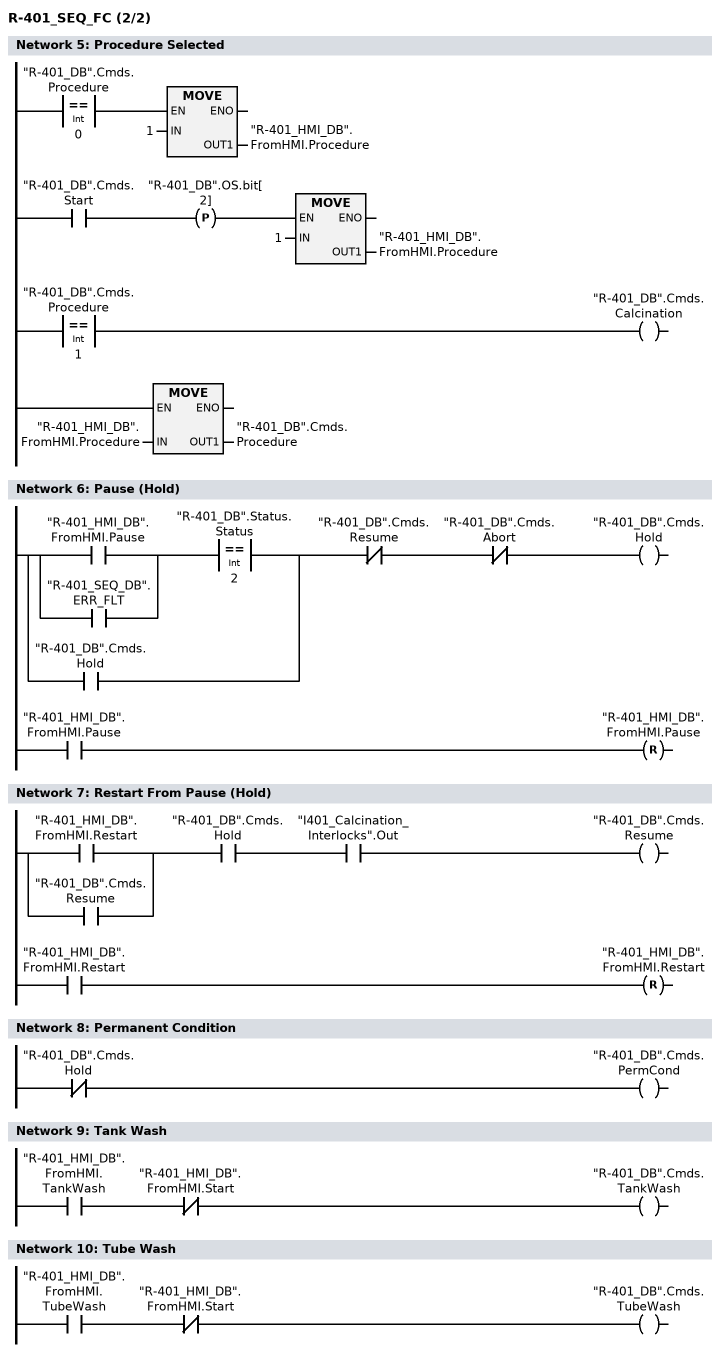
   RUNG wire#powerrail
      { S7_Templates := "SrcType := Int" } EQ_Contact(in1 := "R-401_DB".Cmds.Procedure, in2 := 0)
      Move(in := 1, out1 => "R-401_HMI_DB".FromHMI.Procedure)
   END_RUNG
   RUNG wire#powerrail
      Contact( "R-401_DB".Cmds.Start )
      P_Trig( "R-401_DB".OS.bit[2] )
      Move(in := 1, out1 => "R-401_HMI_DB".FromHMI.Procedure)
   END_RUNG
   RUNG wire#powerrail
      { S7_Templates := "SrcType := Int" } EQ_Contact(in1 := "R-401_DB".Cmds.Procedure, in2 := 1)
      Coil( "R-401_DB".Cmds.Calcination )
   END_RUNG
   RUNG wire#powerrail
      Move(in := "R-401_HMI_DB".FromHMI.Procedure, out1 => "R-401_DB".Cmds.Procedure)
   END_RUNG
   // the same network as SCL:
   IF "R-401_DB".Cmds.Procedure = 0 THEN "R-401_HMI_DB".FromHMI.Procedure := 1; END_IF;
   #_w1 := "R-401_DB".Cmds.Start AND NOT "R-401_DB".OS.bit[2];   // rising edge
   "R-401_DB".OS.bit[2] := "R-401_DB".Cmds.Start;
   IF #_w1 THEN "R-401_HMI_DB".FromHMI.Procedure := 1; END_IF;
   "R-401_DB".Cmds.Calcination := "R-401_DB".Cmds.Procedure = 1;
   "R-401_DB".Cmds.Procedure := "R-401_HMI_DB".FromHMI.Procedure;
END_REGION

REGION Network 6: Pause (Hold)
   RUNG wire#powerrail
      Contact( "R-401_HMI_DB".FromHMI.Pause )
      wire#w1
      { S7_Templates := "SrcType := Int" } EQ_Contact(in1 := "R-401_DB".Status.Status, in2 := 2)
      wire#w2
      I_Contact( "R-401_DB".Cmds.Resume )
      I_Contact( "R-401_DB".Cmds.Abort )
      Coil( "R-401_DB".Cmds.Hold )
   END_RUNG
   RUNG wire#powerrail
      Contact( "R-401_SEQ_DB".ERR_FLT )
   END_RUNG wire#w1
   RUNG wire#powerrail
      Contact( "R-401_DB".Cmds.Hold )
   END_RUNG wire#w2
   RUNG wire#powerrail
      Contact( "R-401_HMI_DB".FromHMI.Pause )
      R_Coil( "R-401_HMI_DB".FromHMI.Pause )
   END_RUNG
   // the same network as SCL:
   "R-401_DB".Cmds.Hold := ((("R-401_HMI_DB".FromHMI.Pause OR "R-401_SEQ_DB".ERR_FLT) AND ("R-401_DB".Status.Status = 2)) OR "R-401_DB".Cmds.Hold) AND NOT "R-401_DB".Cmds.Resume AND NOT "R-401_DB".Cmds.Abort;
   IF "R-401_HMI_DB".FromHMI.Pause THEN "R-401_HMI_DB".FromHMI.Pause := FALSE; END_IF;
END_REGION

REGION Network 7: Restart From Pause (Hold)
   RUNG wire#powerrail
      Contact( "R-401_HMI_DB".FromHMI.Restart )
      wire#w1
      Contact( "R-401_DB".Cmds.Hold )
      Contact( "I401_Calcination_Interlocks".Out )
      Coil( "R-401_DB".Cmds.Resume )
   END_RUNG
   RUNG wire#powerrail
      Contact( "R-401_DB".Cmds.Resume )
   END_RUNG wire#w1
   RUNG wire#powerrail
      Contact( "R-401_HMI_DB".FromHMI.Restart )
      R_Coil( "R-401_HMI_DB".FromHMI.Restart )
   END_RUNG
   // the same network as SCL:
   "R-401_DB".Cmds.Resume := ("R-401_HMI_DB".FromHMI.Restart OR "R-401_DB".Cmds.Resume) AND "R-401_DB".Cmds.Hold AND "I401_Calcination_Interlocks".Out;
   IF "R-401_HMI_DB".FromHMI.Restart THEN "R-401_HMI_DB".FromHMI.Restart := FALSE; END_IF;
END_REGION

REGION Network 8: Permanent Condition
   RUNG wire#powerrail
      I_Contact( "R-401_DB".Cmds.Hold )
      Coil( "R-401_DB".Cmds.PermCond )
   END_RUNG
   // the same network as SCL:
   "R-401_DB".Cmds.PermCond := NOT "R-401_DB".Cmds.Hold;
END_REGION

REGION Network 9: Tank Wash
   RUNG wire#powerrail
      Contact( "R-401_HMI_DB".FromHMI.TankWash )
      I_Contact( "R-401_HMI_DB".FromHMI.Start )
      Coil( "R-401_DB".Cmds.TankWash )
   END_RUNG
   // the same network as SCL:
   "R-401_DB".Cmds.TankWash := "R-401_HMI_DB".FromHMI.TankWash AND NOT "R-401_HMI_DB".FromHMI.Start;
END_REGION

REGION Network 10: Tube Wash
   RUNG wire#powerrail
      Contact( "R-401_HMI_DB".FromHMI.TubeWash )
      I_Contact( "R-401_HMI_DB".FromHMI.Start )
      Coil( "R-401_DB".Cmds.TubeWash )
   END_RUNG
   // the same network as SCL:
   "R-401_DB".Cmds.TubeWash := "R-401_HMI_DB".FromHMI.TubeWash AND NOT "R-401_HMI_DB".FromHMI.Start;
END_REGION

REGION Network 11 (SCL): Sequence Status
   IF "R-401_SEQ_DB".S_NO= 1 THEN
       "R-401_DB".Status.Status := 1; //Idle
   ELSIF (("R-401_SEQ_DB".S_NO > 1 AND "R-401_SEQ_DB".S_NO < 150) OR ("R-401_SEQ_DB".S_NO > 161 AND "R-401_SEQ_DB".S_NO < 170)) AND NOT "R-401_SEQ_DB".ERR_FLT AND NOT "R-401_DB".Cmds.Hold THEN
       "R-401_DB".Status.Status := 2; //Running
   ELSIF "R-401_SEQ_DB".S_NO >= 151 AND "R-401_SEQ_DB".S_NO <= 160 AND NOT "R-401_SEQ_DB".ERR_FLT THEN
       "R-401_DB".Status.Status := 3; // Stopping
   ELSIF  "R-401_SEQ_DB".ERR_FLT AND  (("R-401_SEQ_DB".S_NO > 1 AND "R-401_SEQ_DB".S_NO < 150) OR ("R-401_SEQ_DB".S_NO > 161 AND "R-401_SEQ_DB".S_NO < 170)) THEN
       "R-401_DB".Status.Status := 4; // Held
   ELSIF  "R-401_SEQ_DB".ERR_FLT AND  (("R-401_SEQ_DB".S_NO > 1 AND "R-401_SEQ_DB".S_NO < 150) OR ("R-401_SEQ_DB".S_NO > 161 AND "R-401_SEQ_DB".S_NO < 170)) AND "R-401_Aux_DB"."Bool".TOff  THEN
       "R-401_DB".Status.Status := 5; // Holding
   ELSE
       "R-401_DB".Status.Status := 6; // Unknown
   END_IF;

   "R-401_DB".Status.Running := ("R-401_SEQ_DB".S_NO > 3 AND "R-401_SEQ_DB".S_NO < 150) OR ("R-401_SEQ_DB".S_NO > 161 AND "R-401_SEQ_DB".S_NO < 170);
   "R-401_DB".Status.Initializing := ("R-401_SEQ_DB".S_NO >= 141 AND "R-401_SEQ_DB".S_NO <= 150);

   //Enable/Disable HMI Start/Stop Button
   "R-401_HMI_DB".ToHMI.EnStopButton := ("R-401_DB".Status.Status > 1) OR "R-401_DB".Status.Step = 0; //Enable HMI Stop Button
   "R-401_HMI_DB".ToHMI.EnStartButton := "R-401_DB".Status.Status = 1; //Idle
   "R-401_HMI_DB".ToHMI.EnPauseButton := "R-401_DB".Status.Status = 2; //Enable Pause Button
   "R-401_HMI_DB".ToHMI.EnRestartButton :=  "R-401_DB".Status.Status = 4; //Enable Restart Button

   //****Interlock Activated
   "R-401_HMI_DB".ToHMI.InterlockActivated := "I401_Calcination_Interlocks".Out;
END_REGION

REGION Network 12 (SCL): Sequence Step
   "R-401_DB".Status.Step := "R-401_SEQ_DB".S_NO;
END_REGION

REGION Network 13 (SCL): Sequence state (Procedure running)
   IF "R-401_SEQ_DB".S_NO = 3 OR "R-401_SEQ_DB".S_NO = 4 THEN
       "R-401_DB".Status.State := 1; //Ready
   ELSIF "R-401_SEQ_DB".S_NO >= 21 AND "R-401_SEQ_DB".S_NO <= 60 THEN
       "R-401_DB".Status.State := 2; //Mixing 
   ELSIF "R-401_SEQ_DB".S_NO >= 61 AND "R-401_SEQ_DB".S_NO <= 80 THEN
       "R-401_DB".Status.State := 3; //Pouring
   ELSIF "R-401_SEQ_DB".S_NO >= 141 AND "R-401_SEQ_DB".S_NO <= 150 THEN
       "R-401_DB".Status.State := 4; //Initializing
   ELSIF "R-401_SEQ_DB".S_NO >= 151 AND "R-401_SEQ_DB".S_NO <= 160 THEN
       "R-401_DB".Status.State := 5; //Aborting
   ELSE
       "R-401_DB".Status.State := 0;
   END_IF;
END_REGION

REGION Network 14: Sequence State
END_REGION
END_FUNCTION

FUNCTION "R-401_Tansitions_FC" : Void   // FC98, SCL
{ S7_Optimized_Access := 'TRUE' }
VERSION : 0.1
   VAR_TEMP
      Cond : Struct
         CtrlsOff : Bool;
         Steps : Bool;
      END_STRUCT;
   END_VAR
BEGIN


   //********Controllers Off********
   #Cond.CtrlsOff:= "TC-4011A_R3".MB_Data.Buffer[1] = 0 AND "TC-4011A_R3".MB_Data.Buffer[1] = 0 AND "TC-4011A_R3".MB_Data.Buffer[1] = 0;
   //********Steps********
   #Cond.Steps := "R-401_DB".Status.Step = 25 OR "R-401_DB".Status.Step = 27 OR "R-401_DB".Status.Step = 29;

   //*****************************************Transition conditions**************************************

   "R-401_Aux_DB"."Bool".Cond._001 := #Cond.CtrlsOff;      //"R401_TempMon_DB".ReadyToProcess  AND
END_FUNCTION

// folder: State MACHINE/5)Passivate

FUNCTION "Monitor_R402_FC" : Void   // FC99, LAD
TITLE = FC to call User Functions
{ S7_Optimized_Access := 'TRUE' }
AUTHOR : JL
VERSION : 0.1
BEGIN

REGION Network 1: Moving Furnace temperature to the monitor block
   // Thermocouples:
   // "TT-401A_DB".SAI
   // "TT-401B_DB".SAI
   // "TT-401C_DB".SAI
   // "TT-401C_DB".SAI
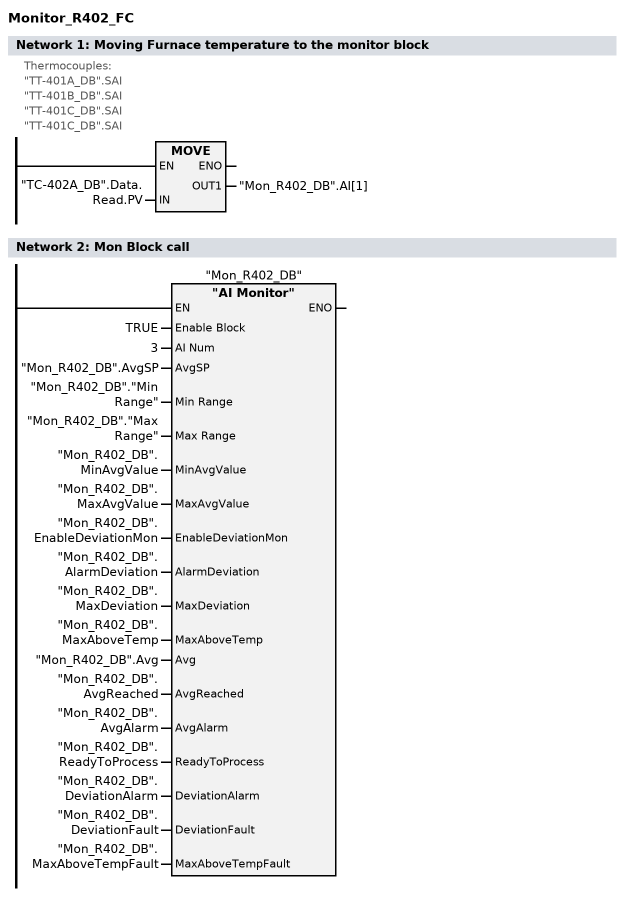
   RUNG wire#powerrail
      Move(in := "TC-402A_DB".Data.Read.PV, out1 => "Mon_R402_DB".AI[1])
   END_RUNG
   // the same network as SCL:
   "Mon_R402_DB".AI[1] := "TC-402A_DB".Data.Read.PV;
END_REGION

REGION Network 2: Mon Block call
   RUNG wire#powerrail
      "Mon_R402_DB"("Enable Block" := TRUE, "AI Num" := 3, AvgSP := "Mon_R402_DB".AvgSP, "Min Range" := "Mon_R402_DB"."Min Range", "Max Range" := "Mon_R402_DB"."Max Range", MinAvgValue := "Mon_R402_DB".MinAvgValue, MaxAvgValue := "Mon_R402_DB".MaxAvgValue, EnableDeviationMon := "Mon_R402_DB".EnableDeviationMon, AlarmDeviation := "Mon_R402_DB".AlarmDeviation, MaxDeviation := "Mon_R402_DB".MaxDeviation, MaxAboveTemp := "Mon_R402_DB".MaxAboveTemp, Avg := "Mon_R402_DB".Avg, AvgReached := "Mon_R402_DB".AvgReached, AvgAlarm := "Mon_R402_DB".AvgAlarm, ReadyToProcess := "Mon_R402_DB".ReadyToProcess, DeviationAlarm := "Mon_R402_DB".DeviationAlarm, DeviationFault := "Mon_R402_DB".DeviationFault, MaxAboveTempFault := "Mon_R402_DB".MaxAboveTempFault)
   END_RUNG
   // the same network as SCL:
   "Mon_R402_DB"("Enable Block" := TRUE,   // "AI Monitor"
                 "AI Num" := 3,
                 AvgSP := "Mon_R402_DB".AvgSP,
                 "Min Range" := "Mon_R402_DB"."Min Range",
                 "Max Range" := "Mon_R402_DB"."Max Range",
                 MinAvgValue := "Mon_R402_DB".MinAvgValue,
                 MaxAvgValue := "Mon_R402_DB".MaxAvgValue,
                 EnableDeviationMon := "Mon_R402_DB".EnableDeviationMon,
                 AlarmDeviation := "Mon_R402_DB".AlarmDeviation,
                 MaxDeviation := "Mon_R402_DB".MaxDeviation,
                 MaxAboveTemp := "Mon_R402_DB".MaxAboveTemp,
                 Avg := "Mon_R402_DB".Avg,
                 AvgReached := "Mon_R402_DB".AvgReached,
                 AvgAlarm := "Mon_R402_DB".AvgAlarm,
                 ReadyToProcess := "Mon_R402_DB".ReadyToProcess,
                 DeviationAlarm := "Mon_R402_DB".DeviationAlarm,
                 DeviationFault := "Mon_R402_DB".DeviationFault,
                 MaxAboveTempFault := "Mon_R402_DB".MaxAboveTempFault);
END_REGION
END_FUNCTION

// folder: State MACHINE/5)Passivate/Reactor R-402

FUNCTION_BLOCK "R-402_SEQ"   // FB31, GRAPH_PLUS
TITLE = Reactor R-401
{ S7_Optimized_Access := 'TRUE' }
AUTHOR : JL
VERSION : 0.1
   VAR_INPUT
      OFF_SQ : Bool := false;   // Turn sequence off
      INIT_SQ : Bool := false;   // Set sequence to initial state
      ACK_EF : Bool := false;   // Acknowledge all errors and faults
      S_PREV : Bool := false;   // Output previous step in parameter S_NO
      S_NEXT : Bool := false;   // Indicate next step in parameter S_NO
      SW_AUTO : Bool := false;   // Automatic mode
      SW_TAP : Bool := false;   // Semiautomatic/switch with transition
      SW_TOP : Bool := false;   // Semiautomatic/ignore transition
      SW_MAN : Bool := false;   // Manual mode
      S_SEL : Int := 0;   // Select step to be output to S_NO
      S_ON : Bool := false;   // Activate step indicated in S_NO
      S_OFF : Bool := false;   // Deactivate step indicated S_NO
      T_PUSH : Bool := false;   // Enable transition to switch in semi automatic mode
   END_VAR
   VAR_OUTPUT
      S_NO : Int := 0;   // Step number
      S_MORE : Bool := false;   // More steps are available and can be shown in S_NO
      S_ACTIVE : Bool := false;   // Step indicated in S_NO is active
      ERR_FLT : Bool := false;   // Interlock or supervision group error
      AUTO_ON : Bool := false;   // Automatic mode is active
      TAP_ON : Bool := false;   // Semiautomatic mode/step with transition enabled
      TOP_ON : Bool := false;   // Semiautomatic mode/ignore transition enabled
      MAN_ON : Bool := false;   // Manual mode is active
   END_VAR
   VAR
      HMI_INFO : Array[0..12] of UInt;
      IF_PAR : G7_IfParPlus_V6;
      RT_DATA : G7_RTDataPlus_V6;   // Internal data area
      Abort : G7_TransitionPlus_V6;   // Transition structure
      InitializeR : G7_TransitionPlus_V6;   // Transition structure
      CalcinP : G7_TransitionPlus_V6;   // Transition structure
      Re : G7_TransitionPlus_V6;   // Transition structure
      Calcinat : G7_TransitionPlus_V6;   // Transition structure
      Wash : G7_TransitionPlus_V6;   // Transition structure
      Shutdwn : G7_TransitionPlus_V6;   // Transition structure
      ColdDDn : G7_TransitionPlus_V6;   // Transition structure
      Std : G7_TransitionPlus_V6;   // Transition structure
      PDn : G7_TransitionPlus_V6;   // Transition structure
      PressRd : G7_TransitionPlus_V6;   // Transition structure
      Rmp1Dn : G7_TransitionPlus_V6;   // Transition structure
      FHldDn : G7_TransitionPlus_V6;   // Transition structure
      Rmp2Dn : G7_TransitionPlus_V6;   // Transition structure
      ScHldDn : G7_TransitionPlus_V6;   // Transition structure
      Rmp3Dn : G7_TransitionPlus_V6;   // Transition structure
      ThHldDn : G7_TransitionPlus_V6;   // Transition structure
      Trans30 : G7_TransitionPlus_V6;   // Transition structure
      Trans31 : G7_TransitionPlus_V6;   // Transition structure
      End : G7_TransitionPlus_V6;   // Transition structure
      Init : G7_TransitionPlus_V6;   // Transition structure
      SAut : G7_TransitionPlus_V6;   // Transition structure
      SIn : G7_TransitionPlus_V6;   // Transition structure
      Initd : G7_TransitionPlus_V6;   // Transition structure
      Ab : G7_TransitionPlus_V6;   // Transition structure
      AbortOn : G7_TransitionPlus_V6;   // Transition structure
      AbortDn : G7_TransitionPlus_V6;   // Transition structure
      ShtSted : G7_TransitionPlus_V6;   // Transition structure
      CldDwnDn : G7_TransitionPlus_V6;   // Transition structure
      DPDn : G7_TransitionPlus_V6;   // Transition structure
      Idle : G7_StepPlus_V6;   // Step structure
      Ready : G7_StepPlus_V6;   // Step structure
      SelectSeq : G7_StepPlus_V6;   // Step structure
      Started : G7_StepPlus_V6;   // Step structure
      "EDIT Params" : G7_StepPlus_V6;   // Step structure
      "USER StartN2" : G7_StepPlus_V6;   // Step structure
      RampUp1 : G7_StepPlus_V6;   // Step structure
      CloseN2 : G7_StepPlus_V6;   // Step structure
      HoldTime : G7_StepPlus_V6;   // Step structure
      SecondHold : G7_StepPlus_V6;   // Step structure
      RampUp3 : G7_StepPlus_V6;   // Step structure
      ThirdHold : G7_StepPlus_V6;   // Step structure
      HeatersOff : G7_StepPlus_V6;   // Step structure
      PressureOff : G7_StepPlus_V6;   // Step structure
      Done : G7_StepPlus_V6;   // Step structure
      Initialize : G7_StepPlus_V6;   // Step structure
      SetAuto : G7_StepPlus_V6;   // Step structure
      SetInitial : G7_StepPlus_V6;   // Step structure
      Initialized : G7_StepPlus_V6;   // Step structure
      AbortStarting : G7_StepPlus_V6;   // Step structure
      Aborting : G7_StepPlus_V6;   // Step structure
      AbortDone : G7_StepPlus_V6;   // Step structure
      ShtdnStarted : G7_StepPlus_V6;   // Step structure
      CoolingDown : G7_StepPlus_V6;   // Step structure
      DePress : G7_StepPlus_V6;   // Step structure
      ShtdnDn : G7_StepPlus_V6;   // Step structure
      SINI : Array[0..5] of USInt;
      LSTT : Array[0..29] of USInt;
      ATAJ : Array[0..29] of USInt;
      ATAB : Array[0..29] of USInt;
      PSTT : Array[0..29] of USInt;
      NSTT : Array[0..29] of USInt;
      ASSJ : Array[0..25] of USInt;
      ASSB : Array[0..25] of USInt;
      PTTS : Array[0..25] of USInt;
      NTTS : Array[0..25] of USInt;
      SW_SQTS : Array[0..25] of USInt;
      SWITCH : Array[0..4] of USInt;
      TVX : Array[0..11] of USInt;
      TTX : Array[0..11] of USInt;
      TSX : Array[0..5] of USInt;
      S00X : Array[0..5] of USInt;
      SOFFX : Array[0..5] of USInt;
      SONX : Array[0..5] of USInt;
      SAX : Array[0..5] of USInt;
      SERRX : Array[0..26] of USInt;
      SMX : Array[0..26] of USInt;
      S0X : Array[0..26] of USInt;
      S1X : Array[0..26] of USInt;
      IL_ALARM_INST : Diag_Alarm;
      SUP_ALARM_INST : Diag_Alarm;
      STEP_TIME_ALARM_INST : Diag_Alarm;
      IEC_TIMER_INST : IEC_TIMER;
      TRANSACTION_FLAG : Bool := false;
   END_VAR
   // SINI[0] := 2;
   // LSTT[0] := 19;
   // NSTT[0] := 19;
   // PTTS[0] := 255;
   // TVX[0] := 16#1;
   // TTX[0] := 16#1;
   // TSX[0] := 16#1;
   // S00X[0] := 16#1;
   // SOFFX[0] := 16#1;
   // SONX[0] := 16#1;
   // SAX[0] := 16#1;
   // SERRX[0] := 16#1;
   // SMX[0] := 16#1;
   // S0X[0] := 16#1;
   // S1X[0] := 16#1;
   // SINI[2] := 255;
   // SINI[3] := 255;
   // SINI[4] := 255;
   // LSTT[1] := 15;
   // LSTT[2] := 255;
   // LSTT[3] := 255;
   // LSTT[4] := 3;
   // LSTT[5] := 255;
   // LSTT[6] := 22;
   // LSTT[16] := 255;
   // LSTT[8] := 255;
   // LSTT[9] := 255;
   // LSTT[10] := 255;
   // LSTT[11] := 255;
   // LSTT[12] := 255;
   // LSTT[13] := 255;
   // LSTT[14] := 255;
   // LSTT[19] := 255;
   // LSTT[22] := 255;
   // LSTT[17] := 255;
   // LSTT[25] := 255;
   // LSTT[20] := 255;
   // LSTT[21] := 255;
   // ATAJ[1] := 1;
   // ATAJ[2] := 2;
   // ATAJ[3] := 3;
   // ATAJ[4] := 4;
   // ATAJ[5] := 5;
   // ATAJ[6] := 6;
   // ATAJ[7] := 7;
   // ATAJ[8] := 8;
   // ATAJ[9] := 9;
   // ATAJ[10] := 10;
   // ATAJ[11] := 11;
   // ATAJ[12] := 12;
   // ATAJ[13] := 13;
   // ATAJ[14] := 14;
   // ATAJ[15] := 15;
   // ATAJ[16] := 16;
   // ATAJ[17] := 17;
   // ATAJ[18] := 18;
   // ATAJ[19] := 19;
   // ATAJ[20] := 20;
   // ATAJ[21] := 21;
   // ATAJ[22] := 22;
   // ATAB[0] := 6;
   // ATAB[1] := 2;
   // ATAB[3] := 3;
   // ATAB[4] := 5;
   // ATAB[5] := 4;
   // ATAB[6] := 1;
   // ATAB[7] := 7;
   // ATAB[8] := 8;
   // ATAB[9] := 9;
   // ATAB[10] := 10;
   // ATAB[11] := 11;
   // ATAB[12] := 12;
   // ATAB[13] := 13;
   // ATAB[14] := 14;
   // ATAB[15] := 15;
   // ATAB[16] := 16;
   // ATAB[17] := 17;
   // ATAB[18] := 18;
   // ATAB[19] := 19;
   // ATAB[20] := 20;
   // ATAB[21] := 21;
   // ATAB[22] := 22;
   // SW_SQTS[21] := 4;
   // SW_SQTS[20] := 4;
   // PSTT[3] := 1;
   // PSTT[4] := 2;
   // PSTT[5] := 2;
   // PSTT[22] := 17;
   // PSTT[7] := 25;
   // PSTT[8] := 3;
   // PSTT[9] := 4;
   // PSTT[10] := 5;
   // PSTT[11] := 6;
   // PSTT[12] := 7;
   // PSTT[13] := 8;
   // PSTT[14] := 9;
   // PSTT[15] := 10;
   // PSTT[16] := 11;
   // PSTT[17] := 13;
   // PSTT[18] := 14;
   // PSTT[19] := 12;
   // PSTT[20] := 15;
   // PSTT[21] := 16;
   // PSTT[25] := 20;
   // NTTS[21] := 26;
   // NTTS[20] := 25;
   // PTTS[21] := 25;
   // PTTS[20] := 24;
   // NSTT[1] := 15;
   // NSTT[2] := 1;
   // NSTT[3] := 2;
   // NSTT[4] := 3;
   // NSTT[5] := 255;
   // NSTT[6] := 22;
   // NSTT[16] := 12;
   // NSTT[8] := 4;
   // NSTT[9] := 5;
   // NSTT[10] := 6;
   // NSTT[11] := 7;
   // NSTT[12] := 8;
   // NSTT[13] := 9;
   // NSTT[14] := 10;
   // NSTT[19] := 13;
   // NSTT[22] := 18;
   // NSTT[17] := 14;
   // NSTT[25] := 21;
   // NSTT[20] := 16;
   // NSTT[21] := 17;
   // ASSJ[20] := 20;
   // ASSB[21] := 21;
   // ASSB[20] := 20;
   // ASSJ[21] := 21;
   // ASSJ[1] := 1;
   // ASSJ[2] := 2;
   // ASSJ[3] := 3;
   // ASSJ[4] := 4;
   // ASSJ[5] := 5;
   // ASSJ[6] := 6;
   // ASSJ[7] := 7;
   // ASSJ[8] := 8;
   // ASSJ[9] := 9;
   // ASSJ[10] := 10;
   // ASSJ[11] := 11;
   // ASSJ[12] := 12;
   // ASSJ[13] := 13;
   // ASSJ[14] := 14;
   // ASSJ[15] := 15;
   // ASSJ[16] := 16;
   // ASSJ[17] := 17;
   // ASSJ[18] := 18;
   // ASSJ[19] := 19;
   // NSTT[23] := 1;
   // NSTT[15] := 11;
   // PSTT[24] := 19;
   // PSTT[23] := 18;
   // ASSB[1] := 1;
   // ASSB[2] := 2;
   // ASSB[3] := 3;
   // ASSB[4] := 4;
   // ASSB[5] := 5;
   // ASSB[6] := 6;
   // ASSB[7] := 7;
   // ASSB[8] := 8;
   // ASSB[9] := 9;
   // ASSB[10] := 10;
   // ASSB[11] := 11;
   // ASSB[12] := 12;
   // ASSB[13] := 13;
   // ASSB[14] := 14;
   // ASSB[15] := 15;
   // ASSB[16] := 16;
   // ASSB[17] := 17;
   // ASSB[18] := 18;
   // ASSB[19] := 19;
   // ATAB[24] := 24;
   // ATAB[23] := 23;
   // ATAJ[24] := 24;
   // ATAJ[23] := 23;
   // PTTS[1] := 2;
   // PTTS[2] := 3;
   // PTTS[3] := 255;
   // PTTS[4] := 8;
   // PTTS[5] := 9;
   // PTTS[6] := 10;
   // PTTS[7] := 11;
   // PTTS[8] := 12;
   // PTTS[9] := 13;
   // PTTS[10] := 14;
   // PTTS[11] := 15;
   // PTTS[12] := 16;
   // PTTS[13] := 19;
   // PTTS[14] := 17;
   // PTTS[15] := 255;
   // PTTS[16] := 20;
   // PTTS[17] := 21;
   // PTTS[18] := 22;
   // PTTS[19] := 255;
   // LSTT[23] := 1;
   // LSTT[15] := 255;
   // NTTS[1] := 3;
   // NTTS[2] := 4;
   // NTTS[3] := 8;
   // NTTS[4] := 9;
   // NTTS[5] := 10;
   // NTTS[6] := 11;
   // NTTS[7] := 12;
   // NTTS[8] := 13;
   // NTTS[9] := 14;
   // NTTS[10] := 15;
   // NTTS[11] := 16;
   // NTTS[12] := 19;
   // NTTS[13] := 17;
   // NTTS[14] := 18;
   // NTTS[15] := 20;
   // NTTS[16] := 21;
   // NTTS[17] := 22;
   // NTTS[18] := 23;
   // NTTS[19] := 24;
   // SW_SQTS[1] := 1;
   // SW_SQTS[2] := 1;
   // SW_SQTS[3] := 2;
   // SW_SQTS[4] := 2;
   // SW_SQTS[5] := 2;
   // SW_SQTS[6] := 2;
   // SW_SQTS[7] := 2;
   // SW_SQTS[8] := 2;
   // SW_SQTS[9] := 2;
   // SW_SQTS[10] := 2;
   // SW_SQTS[11] := 2;
   // SW_SQTS[12] := 2;
   // SW_SQTS[13] := 2;
   // SW_SQTS[14] := 2;
   // SW_SQTS[15] := 3;
   // SW_SQTS[16] := 3;
   // SW_SQTS[17] := 3;
   // SW_SQTS[18] := 3;
   // SW_SQTS[19] := 4;
   // SWITCH[0] := 60;
   // SWITCH[1] := 191;
   // SWITCH[2] := 223;
   // SINI[5] := 255;
   // LSTT[24] := 255;
   // LSTT[28] := 255;
   // LSTT[27] := 255;
   // ATAJ[25] := 25;
   // ATAJ[26] := 26;
   // ATAJ[27] := 27;
   // ATAJ[28] := 28;
   // ATAB[25] := 25;
   // ATAB[26] := 26;
   // ATAB[27] := 27;
   // ATAB[28] := 28;
   // PSTT[26] := 21;
   // PSTT[27] := 22;
   // PSTT[28] := 23;
   // NSTT[24] := 20;
   // NSTT[28] := 24;
   // NSTT[27] := 23;
   // ASSJ[22] := 22;
   // ASSJ[23] := 23;
   // ASSJ[24] := 24;
   // ASSB[22] := 22;
   // ASSB[23] := 23;
   // ASSB[24] := 24;
   // PTTS[22] := 255;
   // PTTS[23] := 27;
   // PTTS[24] := 28;
   // NTTS[22] := 27;
   // NTTS[23] := 28;
   // NTTS[24] := 29;
   // SW_SQTS[22] := 5;
   // SW_SQTS[23] := 5;
   // SW_SQTS[24] := 5;
   // SWITCH[3] := 239;
   // SWITCH[4] := 7;
   // LSTT[29] := 255;
   // ATAJ[29] := 29;
   // ATAB[29] := 29;
   // PSTT[29] := 24;
   // NSTT[29] := 25;
   // ASSJ[25] := 25;
   // ASSB[25] := 25;
   // PTTS[25] := 29;
   // NTTS[25] := 7;
   // SW_SQTS[25] := 5;
BEGIN
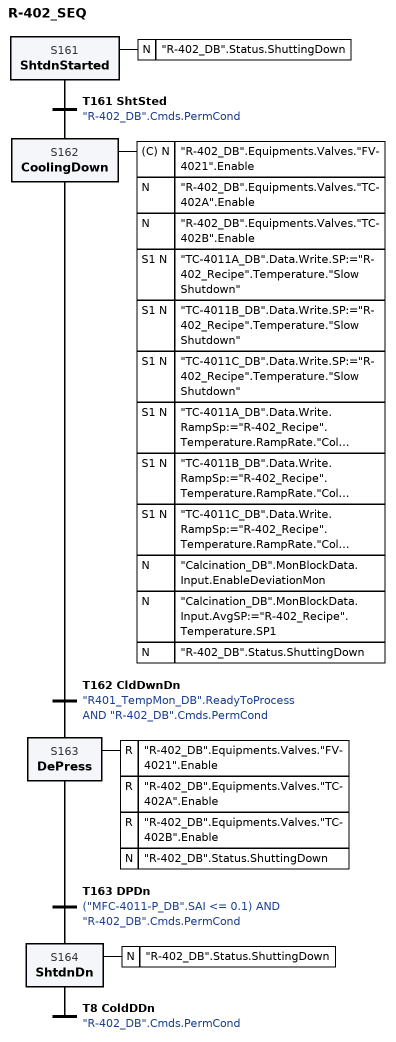
   // permanent pre-instructions
   NETWORK 1
      "R-402_SEQ_FC"();
      "R-402_FC_Inputs"();
      "Monitor_R402_FC"();
      "Alarms"();

   // sequencer 1
   STEP ShtdnStarted:   // S161, max time T#10S, warning time T#7S
      // Shutdown Started
              N    "R-402_DB".Status.ShuttingDown
   END_STEP
   TRANSITION ShtSted FROM ShtdnStarted TO CoolingDown   // T161
      := "R-402_DB".Cmds.PermCond;
   END_TRANSITION
   STEP CoolingDown:   // S162, max time T#10S, warning time T#7S
      (C)     N    "R-402_DB".Equipments.Valves."FV-4021".Enable
              N    "R-402_DB".Equipments.Valves."TC-402A".Enable
              N    "R-402_DB".Equipments.Valves."TC-402B".Enable
          S1  N    "TC-4011A_DB".Data.Write.SP:="R-402_Recipe".Temperature."Slow Shutdown"
          S1  N    "TC-4011B_DB".Data.Write.SP:="R-402_Recipe".Temperature."Slow Shutdown"
          S1  N    "TC-4011C_DB".Data.Write.SP:="R-402_Recipe".Temperature."Slow Shutdown"
          S1  N    "TC-4011A_DB".Data.Write.RampSp:="R-402_Recipe".Temperature.RampRate."Cold Down"
          S1  N    "TC-4011B_DB".Data.Write.RampSp:="R-402_Recipe".Temperature.RampRate."Cold Down"
          S1  N    "TC-4011C_DB".Data.Write.RampSp:="R-402_Recipe".Temperature.RampRate."Cold Down"
              N    "Calcination_DB".MonBlockData.Input.EnableDeviationMon
              N    "Calcination_DB".MonBlockData.Input.AvgSP:="R-402_Recipe".Temperature.SP1
              N    "R-402_DB".Status.ShuttingDown
   END_STEP
   TRANSITION CldDwnDn FROM CoolingDown TO DePress   // T162
      := "R401_TempMon_DB".ReadyToProcess AND "R-402_DB".Cmds.PermCond;
   END_TRANSITION
   STEP DePress:   // S163, max time T#10S, warning time T#7S
              R    "R-402_DB".Equipments.Valves."FV-4021".Enable
              R    "R-402_DB".Equipments.Valves."TC-402A".Enable
              R    "R-402_DB".Equipments.Valves."TC-402B".Enable
              N    "R-402_DB".Status.ShuttingDown
   END_STEP
   TRANSITION DPDn FROM DePress TO ShtdnDn   // T163
      := ("MFC-4011-P_DB".SAI <= 0.1) AND "R-402_DB".Cmds.PermCond;
   END_TRANSITION
   STEP ShtdnDn:   // S164, max time T#10S, warning time T#7S
              N    "R-402_DB".Status.ShuttingDown
   END_STEP
   TRANSITION ColdDDn FROM ShtdnDn TO ?   // T8
      := "R-402_DB".Cmds.PermCond;
   END_TRANSITION

   // permanent post-instructions
   NETWORK 1
      "R-402_FC_Outputs"();
END_FUNCTION_BLOCK

FUNCTION "R-402_FC_Inputs" : Void   // FC94, SCL
{ S7_Optimized_Access := 'TRUE' }
VERSION : 0.1
BEGIN
   //************************************************************************************************************************************
   //************************************************From Eurotherm TC-401A Controllers*********************************************************
   //***************************************************** Working Setpoint (SP)********************************************************
END_FUNCTION

FUNCTION "R-402_FC_Outputs" : Void   // FC95, SCL
{ S7_Optimized_Access := 'TRUE' }
VERSION : 0.1
   VAR_TEMP
      XV : Struct
         "4021" : Bool;
         "4022" : Bool;
         "4024" : Bool;
         "4025" : Bool;
      END_STRUCT;
      "FV-4021" : Struct
         On : Bool;
         Cond_1 : Bool;
      END_STRUCT;
      "FV-4024" : Struct
         On : Bool;
         Cond_1 : Bool;
      END_STRUCT;
      "FV-4025" : Struct
         On : Bool;
         Cond_1 : Bool;
      END_STRUCT;
      "TC-402A" : Struct
         On : Bool;
         Cond_1 : Bool;
      END_STRUCT;
      "TC-402B" : Struct
         On : Bool;
         Cond_1 : Bool;
      END_STRUCT;
   END_VAR
BEGIN
   //****** Equipmens Activation*******
   //
   //**************************************************************
   //
   //***********************************************H2 Inlet Furnace Valve**********************************************************************
   IF "XV-4021_DB".Mode = 0 THEN
       "R-402_DB".Equipments.Valves."XV-4021".CmdOn := "R-402_DB".Equipments.Valves."XV-4021".Enable AND NOT "R-402_DB".Cmds.Hold AND NOT "R-402_DB".Status.Aborting;
       //Delay Off To avoid Overpressure the Lines
       #XV."4021" := "R-402_DB".Equipments.Valves."XV-4021".CmdOn;
       "R-402_Aux_DB".Timer."XV-4021".TOF(IN := #XV."4021",
       PT := "R-402_Aux_DB".Constants.CmdDelay);
       //Command to the Valve
       IF "R-402_Aux_DB".Timer."XV-4021".Q THEN
           "XV-4021_DB".CMD := 2;
       ELSE
           "XV-4021_DB".CMD := 1;
       END_IF;
       "R-402_DB".Equipments.Valves."XV-4021".TurningOff := NOT "R-402_DB".Equipments.Valves."XV-4021".CmdOn AND "R-402_Aux_DB".Timer."XV-4021".Q;
   END_IF;
   //***********************************************N2 (Second)Inlet Furnace Valve**********************************************************************
   IF "XV-4022_DB".Mode = 0 THEN
       "R-402_DB".Equipments.Valves."XV-4022".CmdOn := "R-402_DB".Equipments.Valves."XV-4022".Enable AND NOT "R-402_DB".Cmds.Hold AND NOT "R-402_DB".Status.Aborting;
       //Delay Off To avoid Overpressure the Lines
       #XV."4022" := "R-402_DB".Equipments.Valves."XV-4022".CmdOn;
       "R-402_Aux_DB".Timer."XV-4022".TOF(IN := #XV."4022",
                                          PT := "R-402_Aux_DB".Constants.CmdDelay);
       //Command to the Valve
       IF "R-402_Aux_DB".Timer."XV-4022".Q THEN
           "XV-4022_DB".CMD := 2;
       ELSE
           "XV-4022_DB".CMD := 1;
       END_IF;
       "R-402_DB".Equipments.Valves."XV-4022".TurningOff := NOT "R-402_DB".Equipments.Valves."XV-4022".CmdOn AND "R-402_Aux_DB".Timer."XV-4022".Q;
   END_IF;
   //***********************************************Air Inlet Furnace Valve**********************************************************************
   IF "XV-4024_DB".Mode = 0 THEN
       "R-402_DB".Equipments.Valves."XV-4024".CmdOn := "R-402_DB".Equipments.Valves."XV-4024".Enable AND NOT "R-402_DB".Cmds.Hold AND NOT "R-402_DB".Status.Aborting;
       //Delay Off To avoid Overpressure the Lines
       #XV."4024" := "R-402_DB".Equipments.Valves."XV-4024".CmdOn;
       "R-402_Aux_DB".Timer."XV-4024".TOF(IN := #XV."4024",
                                          PT := "R-402_Aux_DB".Constants.CmdDelay);
       //Command to the Valve
       IF "R-402_Aux_DB".Timer."XV-4024".Q THEN
           "XV-4024_DB".CMD := 2;
       ELSE
           "XV-4024_DB".CMD := 1;
       END_IF;
       "R-402_DB".Equipments.Valves."XV-4024".TurningOff := NOT "R-402_DB".Equipments.Valves."XV-4024".CmdOn AND "R-402_Aux_DB".Timer."XV-4024".Q; 
   END_IF;
   //***********************************************N2 (First)Inlet Furnace Valve**********************************************************************
   IF "XV-4025_DB".Mode = 0 THEN
       "R-402_DB".Equipments.Valves."XV-4025".CmdOn := "R-402_DB".Equipments.Valves."XV-4025".Enable AND NOT "R-402_DB".Cmds.Hold AND NOT "R-402_DB".Status.Aborting;
       //Delay Off To avoid Overpressure the Lines
       #XV."4025" := "R-402_DB".Equipments.Valves."XV-4025".CmdOn;
       "R-402_Aux_DB".Timer."XV-4025".TOF(IN := #XV."4025",
                                          PT := "R-402_Aux_DB".Constants.CmdDelay);
       //Command to the Valve
       IF "R-402_Aux_DB".Timer."XV-4025".Q THEN
           "XV-4025_DB".CMD := 2;
       ELSE
           "XV-4025_DB".CMD := 1;
       END_IF;
       "R-402_DB".Equipments.Valves."XV-4025".TurningOff := NOT "R-402_DB".Equipments.Valves."XV-4025".CmdOn AND "R-402_Aux_DB".Timer."XV-4025".Q;
   END_IF;

   //**********************************TC-402A  Temperature Control (TIC-402A)**************************************************
   #"TC-402A".Cond_1 := "R-402_DB".Equipments.Valves."TC-402A".Enable AND NOT "R-402_Aux_DB".Timer.HoldTimer.Q;
   "R-402_DB".Equipments.Valves."TC-402A".CmdOn := #"TC-402A".Cond_1 AND NOT "R-402_DB".Cmds.Hold AND NOT "R-402_DB".Status.Aborting;
   //On Command to the Controller
   #"TC-402A".On := "R-402_DB".Equipments.Valves."TC-402A".CmdOn;

   IF #"TC-402A".On  THEN 
       "TIC-R402A_DB".enableManualMode := False;
       "TIC-R402A_DB".enableRemoteSetpoint := False;
       "TIC-R402A_DB".hmi.Controls.manualEnable := False;
       "TIC-R402A_DB".hmi.Config.mode := 3;

       "TC-R402A_Ramp_DB".Enable := TRUE;    //Enable the Ramp function.
   ELSE
       "TC-R402A_Ramp_DB".Enable := FALSE;


   END_IF;

   //**********************************TC-402B Temperature Control (TIC-402B)**************************************************
   #"TC-402B".Cond_1 := "R-402_DB".Equipments.Valves."TC-402B".Enable AND NOT "R-402_Aux_DB".Timer.HoldTimer.Q;
   "R-402_DB".Equipments.Valves."TC-402B".CmdOn := #"TC-402B".Cond_1 AND NOT "R-402_DB".Cmds.Hold AND NOT "R-402_DB".Status.Aborting;
   //On Command to the Controller
   #"TC-402B".On := "R-402_DB".Equipments.Valves."TC-402B".CmdOn;

   IF #"TC-402B".On THEN
       "TIC-R402B_DB".enableManualMode := False;
       "TIC-R402B_DB".enableRemoteSetpoint := False;
       "TIC-R402B_DB".hmi.Controls.manualEnable := False;
       "TIC-R402B_DB".hmi.Config.mode := 3;

       "TC-R402B_Ramp_DB".Enable := TRUE;    //Enable the Ramp function.
   ELSE
       "TC-R402B_Ramp_DB".Enable := FALSE;


   END_IF;

   //**********************************FV-4021 H2 Flow Control Valve (MFC-4021)******************************************************
   IF "FV-4021_DB".HMI.Config.Mode = 0 THEN
       #"FV-4021".Cond_1 := "R-402_DB".Equipments.Valves."FV-4021".Enable;
       "R-402_DB".Equipments.Valves."FV-4021".CmdOn := #"FV-4021".Cond_1 AND NOT "R-402_DB".Cmds.Hold AND NOT "R-402_DB".Status.Aborting;
       //Delay Off To avoid Overpressure the Lines
       #"FV-4021".On := "R-402_DB".Equipments.Valves."FV-4021".CmdOn;
       "R-402_Aux_DB".Timer."FV-4021".TOF(IN := #"FV-4021".On,
                                          PT := "R-402_Aux_DB".Constants.CmdDelay);
       IF "R-402_Aux_DB".Timer."FV-4021".Q THEN

           // "MFC-4021_DB_MB".Data.SP := "R-402_Recipe".Reduction."H2 Flow SP";

           "MFC-4021_DB".enableManualMode := False;
           "MFC-4021_DB".enableRemoteSetpoint := False;
           "MFC-4021_DB".hmi.Controls.manualEnable := False;
           "MFC-4021_DB".hmi.Config.mode := 3;
       END_IF;//  ELSE
         //  "MFC-4021_DB".enableManualMode := True;
         //  "MFC-4021_DB".hmi.Controls.manualEnable := True;
         //  "MFC-4021_DB".hmi.Config.mode := 4;
          // "MFC-4021_DB".hmi.Controls.manualOutput := "R-402_Recipe".Reduction.Shutdown;

          // "MFC-4021_DB_MB".Data.SP := "R-402_Recipe".Reduction.Shutdown;

      // END_IF;
       "R-402_DB".Equipments.Valves."FV-4021".TurningOff := NOT "R-402_DB".Equipments.Valves."FV-4021".CmdOn AND "R-402_Aux_DB".Timer."XV-4021".Q;
   END_IF;

   //**********************************FV-4024 Air Pressure Control Valve (MFC-4024)******************************************************
   IF "FV-4024_DB".HMI.Config.Mode = 0 THEN
       #"FV-4024".Cond_1 := "R-402_DB".Equipments.Valves."FV-4024".Enable;
       "R-402_DB".Equipments.Valves."FV-4024".CmdOn := #"FV-4024".Cond_1 AND NOT "R-402_DB".Cmds.Hold AND NOT "R-402_DB".Status.Aborting;
       //Delay Off To avoid Overpressure the Lines
       #"FV-4024".On := "R-402_DB".Equipments.Valves."FV-4024".CmdOn;
       "R-402_Aux_DB".Timer."FV-4024".TOF(IN := #"FV-4024".On,
                                          PT := "R-402_Aux_DB".Constants.CmdDelay);
       IF "R-402_Aux_DB".Timer."FV-4024".Q THEN

           // "MFC-4024_DB_MB".Data.SP := "R-402_Recipe".Reduction."Air pressure SP";

           "MFC-4024_DB".enableManualMode := False;
           "MFC-4024_DB".enableRemoteSetpoint := False;
           "MFC-4024_DB".hmi.Controls.manualEnable := False;
           "MFC-4024_DB".hmi.Config.mode := 3;
       END_IF;//    ELSE
          // "MFC-4024_DB_MB".Data.SP := "R-402_Recipe".Reduction.Shutdown;

         //  "MFC-4024_DB".enableManualMode := True;
         //  "MFC-4024_DB".hmi.Controls.manualEnable := True;
         //  "MFC-4024_DB".hmi.Config.mode := 4;
          // "MFC-4024_DB".hmi.Controls.manualOutput := "R-402_Recipe".Reduction.Shutdown;

     //  END_IF;
       "R-402_DB".Equipments.Valves."FV-4024".TurningOff := NOT "R-402_DB".Equipments.Valves."FV-4024".CmdOn AND "R-402_Aux_DB".Timer."XV-4024".Q;
   END_IF;

   //**********************************FV-4025 N2 Pressure Control Valve (MFC-4025)******************************************************
   IF "FV-4025_DB".HMI.Config.Mode = 0 THEN
       #"FV-4025".Cond_1 := "R-402_DB".Equipments.Valves."FV-4025".Enable;
       "R-402_DB".Equipments.Valves."FV-4025".CmdOn := #"FV-4025".Cond_1 AND NOT "R-402_DB".Cmds.Hold AND NOT "R-402_DB".Status.Aborting;
       //Delay Off To avoid Overpressure the Lines
       #"FV-4025".On := "R-402_DB".Equipments.Valves."FV-4025".CmdOn;
       "R-402_Aux_DB".Timer."FV-4025".TOF(IN := #"FV-4025".On,
                                          PT := "R-402_Aux_DB".Constants.CmdDelay);
       IF "R-402_Aux_DB".Timer."FV-4025".Q THEN

           // "MFC-4025_DB_MB".Data.SP := "R-402_Recipe".Reduction."N2 Pressure SP";

           "MFC-4025_DB".enableManualMode := False;
           "MFC-4025_DB".enableRemoteSetpoint := False;
           "MFC-4025_DB".hmi.Controls.manualEnable := False;
           "MFC-4025_DB".hmi.Config.mode := 3;
       END_IF; // ELSE
          // "MFC-4025_DB_MB".Data.SP := "R-402_Recipe".Reduction.Shutdown;

          // "MFC-4025_DB".enableManualMode := True;
         //  "MFC-4025_DB".hmi.Controls.manualEnable := True;
         //  "MFC-4025_DB".hmi.Config.mode := 4;
        //   "MFC-4025_DB".hmi.Controls.manualOutput := "R-402_Recipe".Reduction.Shutdown;

     //  END_IF;
       "R-402_DB".Equipments.Valves."FV-4025".TurningOff := NOT "R-402_DB".Equipments.Valves."FV-4025".CmdOn AND "R-402_Aux_DB".Timer."XV-4025".Q;
   END_IF;

   //******************************************************************************************************************************************//
   //**************************************************To Temperature Controllers**************************************************************




       //**********ALICAT Controllers************//
       //***********************************************ALICAT Control Selection*******************************************************//
       //Command ID and Command Argument 
       (*With this Values the Selection is:
           Address 1000=11; Change control loop variable
           Address 1001=3;  Absolute Pressure*)
   //******************H2 Flow Controll3er******************************************
   "MFC-4021_MB_WCMD_DB".MB_Data.Buffer[1] := 11;
   "MFC-4021_MB_WCMD_DB".MB_Data.Buffer[2] := 3;
   //******************Air Flow Controll3er******************************************
   "MFC-4024_MB_WCMD_DB".MB_Data.Buffer[1] := 11;
   "MFC-4024_MB_WCMD_DB".MB_Data.Buffer[2] := 3;
   //*******************N2 Flow Controll3er******************************************
   "MFC-4025_MB_WCMD_DB".MB_Data.Buffer[1] := 11;
   "MFC-4025_MB_WCMD_DB".MB_Data.Buffer[2] := 3;
    //***********************************************ALICAT Controller Set Point*******************************************************//
   //"MFC-4021_MB_W_DB".MB_Data.Buffer[1] := "MFC-4021_DB_MB".Data.SP;
   //"MFC-4024_MB_W_DB".MB_Data.Buffer[1] := "MFC-4024_DB_MB".Data.SP;
   //"MFC-4025_MB_W_DB".MB_Data.Buffer[1] := "MFC-4025_DB_MB".Data.SP;
   //*********MFC-4021*******
   "MFC-4021_MB_W_DB".MB_Data.Buffer[1] := (INT_TO_REAL("FV-4021_DB".CMD) * 100) / 27648.0;
   "MFC-4021_DB_MB".Data.SP := "MFC-4021_MB_W_DB".MB_Data.Buffer[1];
   //*********MFC-4024*******
   "MFC-4024_MB_W_DB".MB_Data.Buffer[1] := (INT_TO_REAL("FV-4024_DB".CMD) * 100) / 27648.0;
   "MFC-4024_DB_MB".Data.SP := "MFC-4024_MB_W_DB".MB_Data.Buffer[1];
   //*********MFC-4025*******
   "MFC-4025_MB_W_DB".MB_Data.Buffer[1] := (INT_TO_REAL("FV-4025_DB".CMD) * 100) / 27648.0;
   "MFC-4025_DB_MB".Data.SP := "MFC-4025_MB_W_DB".MB_Data.Buffer[1];